(* Logix 5000 project; controller FV vendor 1 type 14 code 217 rev 31.11; software revision 31.00; part 42 of 63 *)
(* tags used below, declared in another part *)
   FV_B100 : INT[255];   // FV FLAGS
   FV_B100_0_1_OutputBit : BOOL;
   FV_N101 : INT[255];   // FV INT Fermentation control integer workspace
   FV_N110 : INT[255];   // FV DATA 0 CURRENT FV DATA
   FV_N12 : INT[255];   // SYS_PARMS System Parameter Fil e
   FV_SFile : INT[255];   // SLC Equivalent System File, So Original Code Can Remain
   FV_T102 : TIMER[20];
   FV_T4 : TIMER[10];
(* FV_Common, continued *)

ROUTINE FV_FV_ELAPSED_102   (* ladder *)
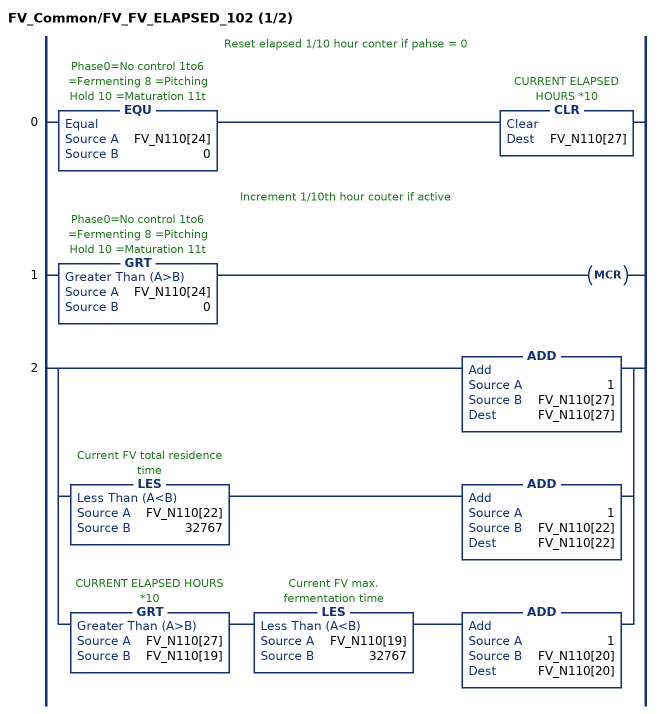
   // Reset elapsed 1/10 hour conter if pahse = 0
   0: EQU(FV_N110[24],0)CLR(FV_N110[27]);
   // Increment 1/10th hour couter if active
   1: GRT(FV_N110[24],0)MCR();
   2: [ADD(1,FV_N110[27],FV_N110[27]) ,LES(FV_N110[22],32767) ADD(1,FV_N110[22],FV_N110[22]) ,GRT(FV_N110[27],FV_N110[19]) LES(FV_N110[19],32767) ADD(1,FV_N110[20],FV_N110[20]) ];
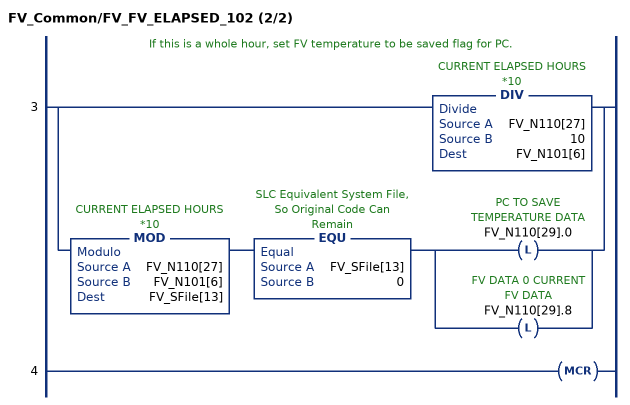
   // If this is a whole hour, set FV temperature to be saved flag for PC.
   3: [DIV(FV_N110[27],10,FV_N101[6]) ,MOD(FV_N110[27],FV_N101[6],FV_SFile[13]) EQU(FV_SFile[13],0) [OTL(FV_N110[29].0) ,OTL(FV_N110[29].8) ] ];
   4: MCR();
END_ROUTINE

ROUTINE FV_FV_MCP_100   (* ladder *)
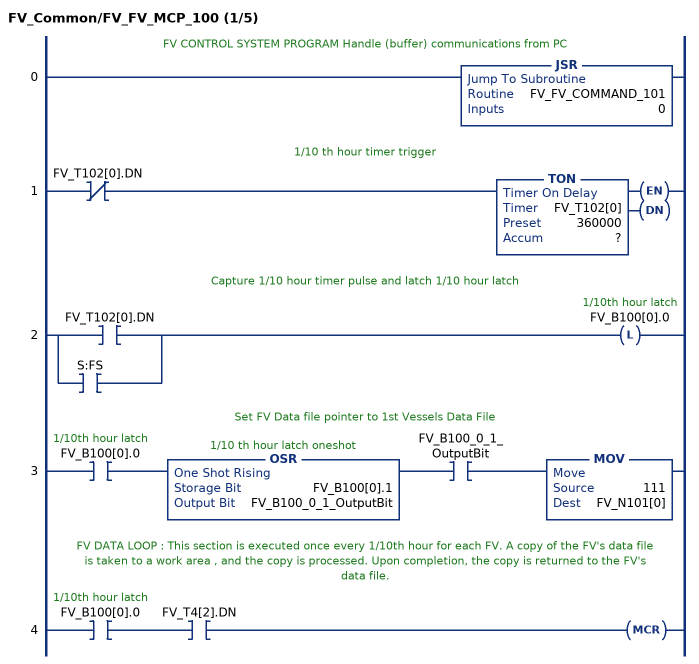
   // FV CONTROL SYSTEM PROGRAM Handle (buffer) communications from PC
   0: JSR(FV_FV_COMMAND_101,0);
   // 1/10 th hour timer trigger
   1: XIO(FV_T102[0].DN)TON(FV_T102[0],?,?);
   // Capture 1/10 hour timer pulse and latch 1/10 hour latch
   2: [XIC(FV_T102[0].DN) ,XIC(S:FS) ]OTL(FV_B100[0].0);
   // Set FV Data file pointer to 1st Vessels Data File
   3: XIC(FV_B100[0].0)OSR(FV_B100[0].1,FV_B100_0_1_OutputBit)XIC(FV_B100_0_1_OutputBit)MOV(111,FV_N101[0]);
   // FV DATA LOOP : This section is executed once every 1/10th hour for each FV. A copy of the FV's data file is taken to a work area , and the copy is processed. Upon completion, the copy is returned to the FV's data file.
   4: XIC(FV_B100[0].0)XIC(FV_T4[2].DN)MCR();
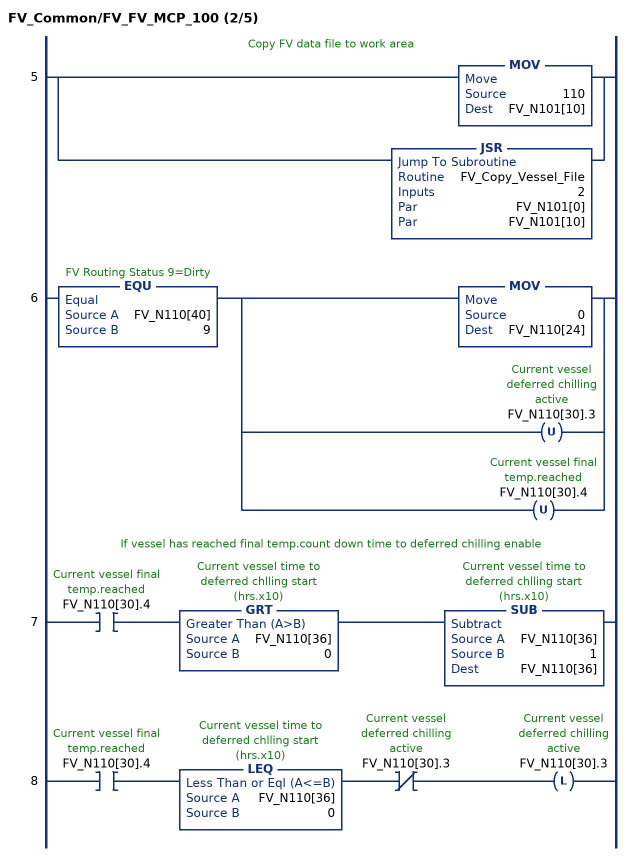
   // Copy FV data file to work area
   5: [MOV(110,FV_N101[10]) ,JSR(FV_Copy_Vessel_File,2,FV_N101[0],FV_N101[10]) ];
   6: EQU(FV_N110[40],9)[MOV(0,FV_N110[24]) ,OTU(FV_N110[30].3) ,OTU(FV_N110[30].4) ];
   // If vessel has reached final temp.count down time to deferred chilling enable
   7: XIC(FV_N110[30].4)GRT(FV_N110[36],0)SUB(FV_N110[36],1,FV_N110[36]);
   8: XIC(FV_N110[30].4)LEQ(FV_N110[36],0)XIO(FV_N110[30].3)OTL(FV_N110[30].3);
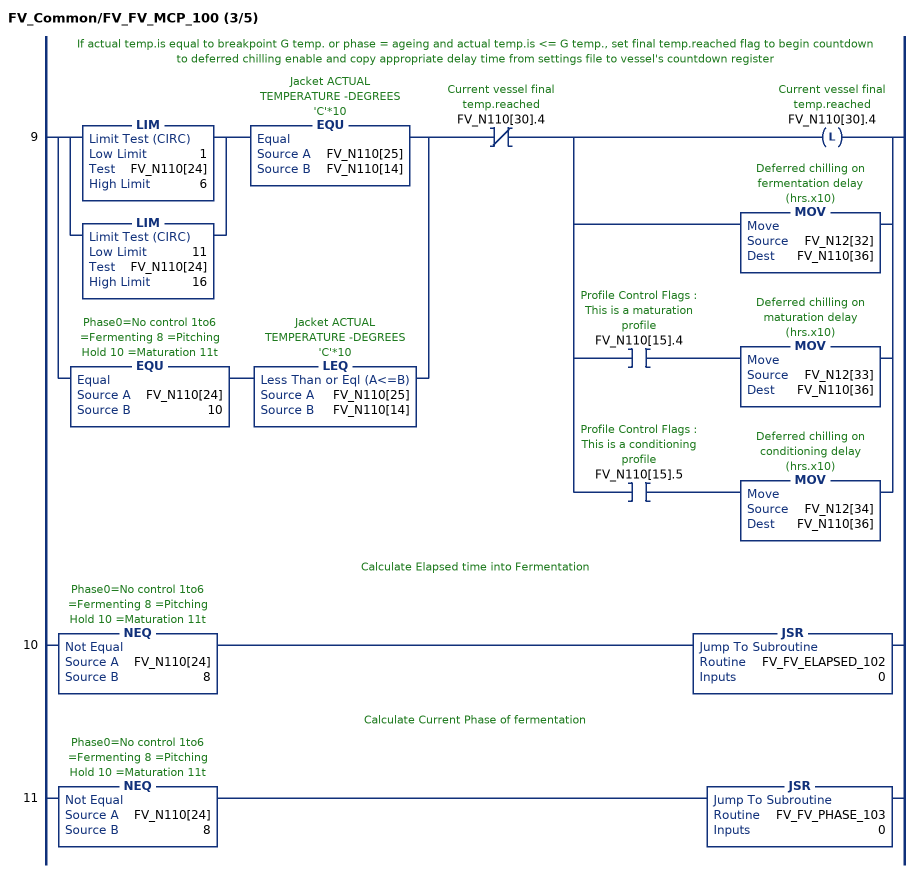
   // If actual temp.is equal to breakpoint G temp. or phase = ageing and actual temp.is <= G temp., set final temp.reached flag to begin countdown to deferred chilling enable and copy appropriate delay time from settings file to vessel's countdown register
   9: [[LIM(1,FV_N110[24],6) ,LIM(11,FV_N110[24],16) ] EQU(FV_N110[25],FV_N110[14]) ,EQU(FV_N110[24],10) LEQ(FV_N110[25],FV_N110[14]) ]XIO(FV_N110[30].4)[OTL(FV_N110[30].4) ,MOV(FV_N12[32],FV_N110[36]) ,XIC(FV_N110[15].4) MOV(FV_N12[33],FV_N110[36]) ,XIC(FV_N110[15].5) MOV(FV_N12[34],FV_N110[36]) ];
   // Calculate Elapsed time into Fermentation
   10: NEQ(FV_N110[24],8)JSR(FV_FV_ELAPSED_102,0);
   // Calculate Current Phase of fermentation
   11: NEQ(FV_N110[24],8)JSR(FV_FV_PHASE_103,0);
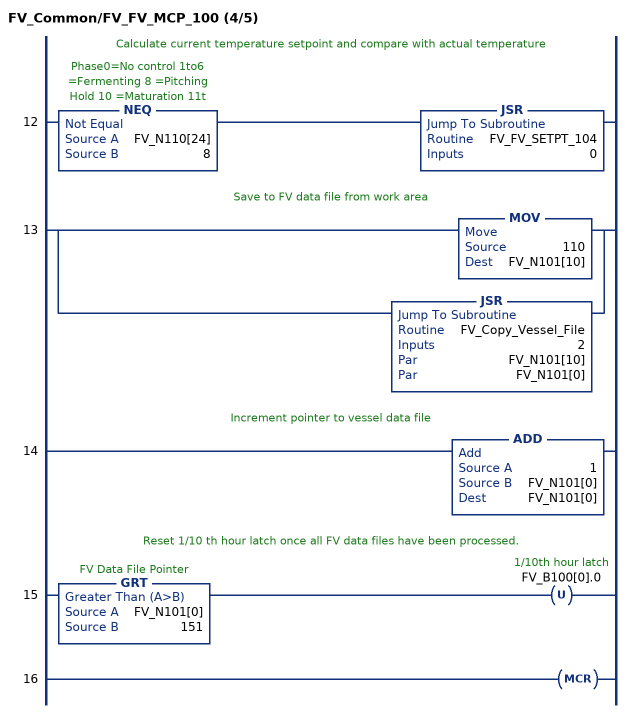
   // Calculate current temperature setpoint and compare with actual temperature
   12: NEQ(FV_N110[24],8)JSR(FV_FV_SETPT_104,0);
   // Save to FV data file from work area
   13: [MOV(110,FV_N101[10]) ,JSR(FV_Copy_Vessel_File,2,FV_N101[10],FV_N101[0]) ];
   // Increment pointer to vessel data file
   14: ADD(1,FV_N101[0],FV_N101[0]);
   // Reset 1/10 th hour latch once all FV data files have been processed.
   15: GRT(FV_N101[0],151)OTU(FV_B100[0].0);
   16: MCR();
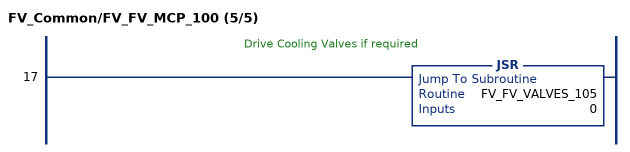
   // Drive Cooling Valves if required
   17: JSR(FV_FV_VALVES_105,0);
END_ROUTINE

ROUTINE FV_FV_PHASE_103   (* ladder *)
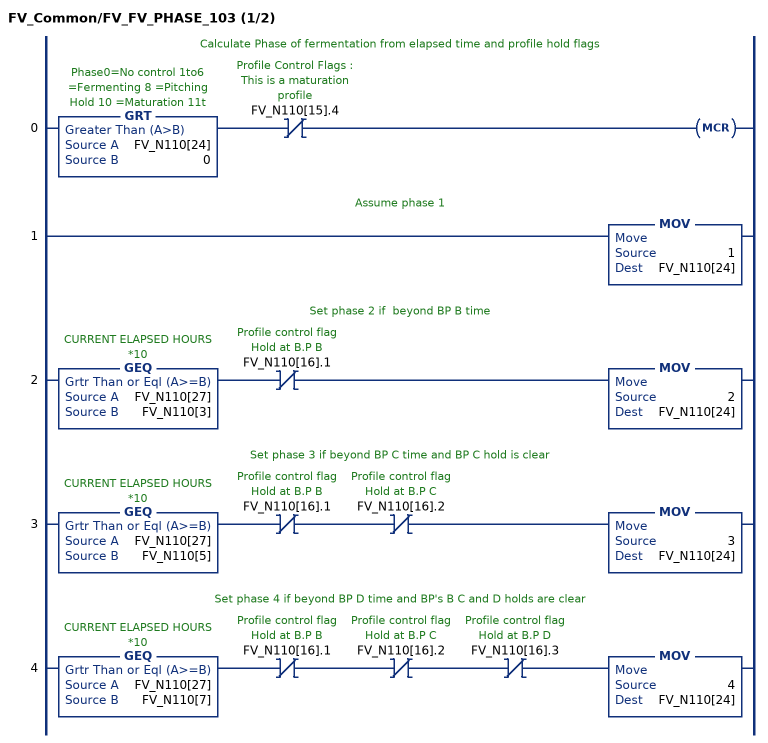
   // Calculate Phase of fermentation from elapsed time and profile hold flags
   0: GRT(FV_N110[24],0)XIO(FV_N110[15].4)MCR();
   // Assume phase 1
   1: MOV(1,FV_N110[24]);
   // Set phase 2 if  beyond BP B time
   2: GEQ(FV_N110[27],FV_N110[3])XIO(FV_N110[16].1)MOV(2,FV_N110[24]);
   // Set phase 3 if beyond BP C time and BP C hold is clear
   3: GEQ(FV_N110[27],FV_N110[5])XIO(FV_N110[16].1)XIO(FV_N110[16].2)MOV(3,FV_N110[24]);
   // Set phase 4 if beyond BP D time and BP's B C and D holds are clear
   4: GEQ(FV_N110[27],FV_N110[7])XIO(FV_N110[16].1)XIO(FV_N110[16].2)XIO(FV_N110[16].3)MOV(4,FV_N110[24]);
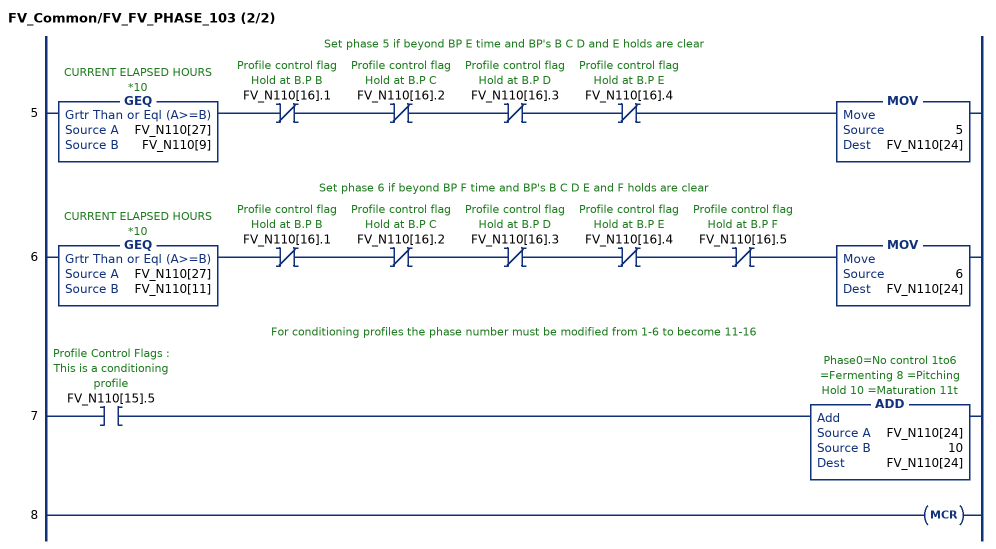
   // Set phase 5 if beyond BP E time and BP's B C D and E holds are clear
   5: GEQ(FV_N110[27],FV_N110[9])XIO(FV_N110[16].1)XIO(FV_N110[16].2)XIO(FV_N110[16].3)XIO(FV_N110[16].4)MOV(5,FV_N110[24]);
   // Set phase 6 if beyond BP F time and BP's B C D E and F holds are clear
   6: GEQ(FV_N110[27],FV_N110[11])XIO(FV_N110[16].1)XIO(FV_N110[16].2)XIO(FV_N110[16].3)XIO(FV_N110[16].4)XIO(FV_N110[16].5)MOV(6,FV_N110[24]);
   // For conditioning profiles the phase number must be modified from 1-6 to become 11-16
   7: XIC(FV_N110[15].5)ADD(FV_N110[24],10,FV_N110[24]);
   8: MCR();
END_ROUTINE

ROUTINE FV_FV_SETPT_104   (* ladder *)
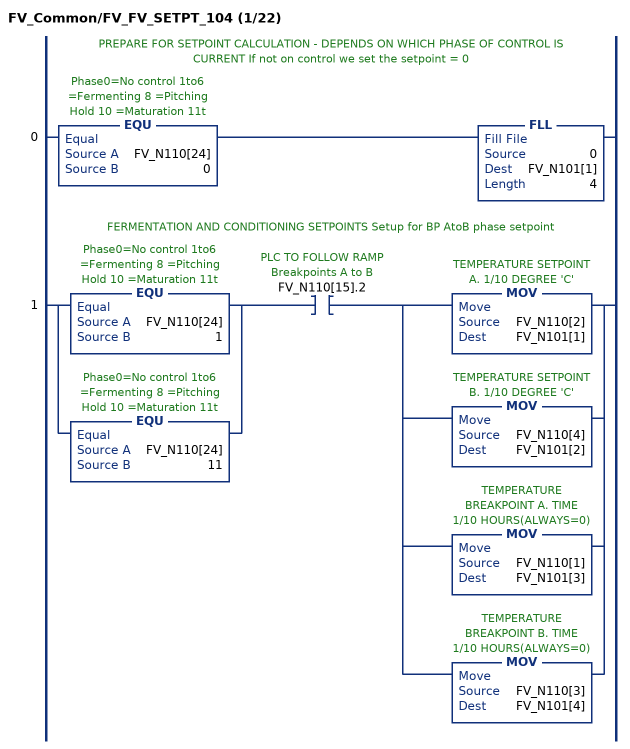
   // PREPARE FOR SETPOINT CALCULATION - DEPENDS ON WHICH PHASE OF CONTROL IS CURRENT If not on control we set the setpoint = 0
   0: EQU(FV_N110[24],0)FLL(0,FV_N101[1],4);
   // FERMENTATION AND CONDITIONING SETPOINTS Setup for BP AtoB phase setpoint
   1: [EQU(FV_N110[24],1) ,EQU(FV_N110[24],11) ]XIC(FV_N110[15].2)[MOV(FV_N110[2],FV_N101[1]) ,MOV(FV_N110[4],FV_N101[2]) ,MOV(FV_N110[1],FV_N101[3]) ,MOV(FV_N110[3],FV_N101[4]) ];
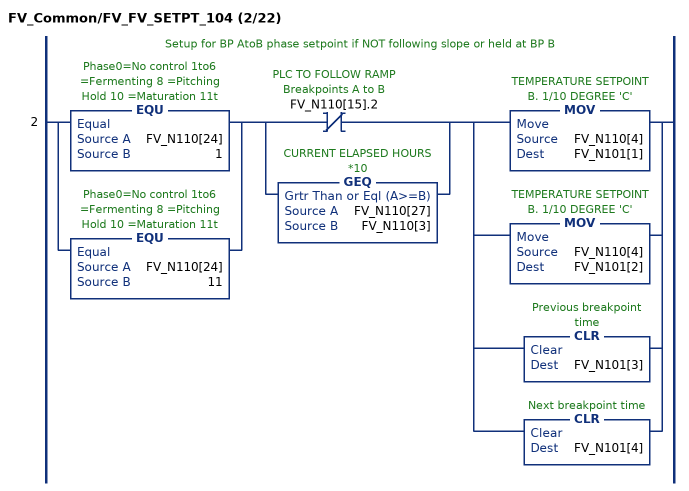
   // Setup for BP AtoB phase setpoint if NOT following slope or held at BP B
   2: [EQU(FV_N110[24],1) ,EQU(FV_N110[24],11) ][XIO(FV_N110[15].2) ,GEQ(FV_N110[27],FV_N110[3]) ][MOV(FV_N110[4],FV_N101[1]) ,MOV(FV_N110[4],FV_N101[2]) ,CLR(FV_N101[3]) ,CLR(FV_N101[4]) ];
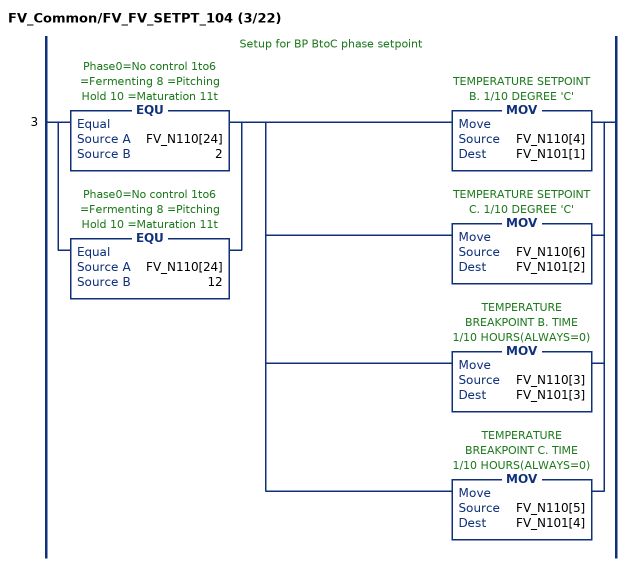
   // Setup for BP BtoC phase setpoint
   3: [EQU(FV_N110[24],2) ,EQU(FV_N110[24],12) ][MOV(FV_N110[4],FV_N101[1]) ,MOV(FV_N110[6],FV_N101[2]) ,MOV(FV_N110[3],FV_N101[3]) ,MOV(FV_N110[5],FV_N101[4]) ];
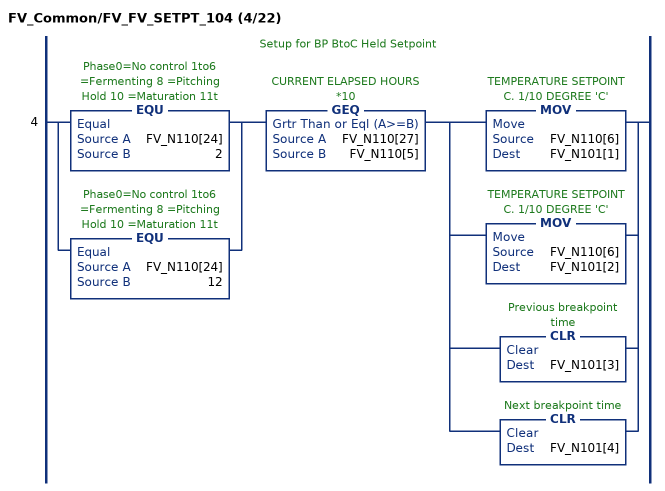
   // Setup for BP BtoC Held Setpoint
   4: [EQU(FV_N110[24],2) ,EQU(FV_N110[24],12) ]GEQ(FV_N110[27],FV_N110[5])[MOV(FV_N110[6],FV_N101[1]) ,MOV(FV_N110[6],FV_N101[2]) ,CLR(FV_N101[3]) ,CLR(FV_N101[4]) ];
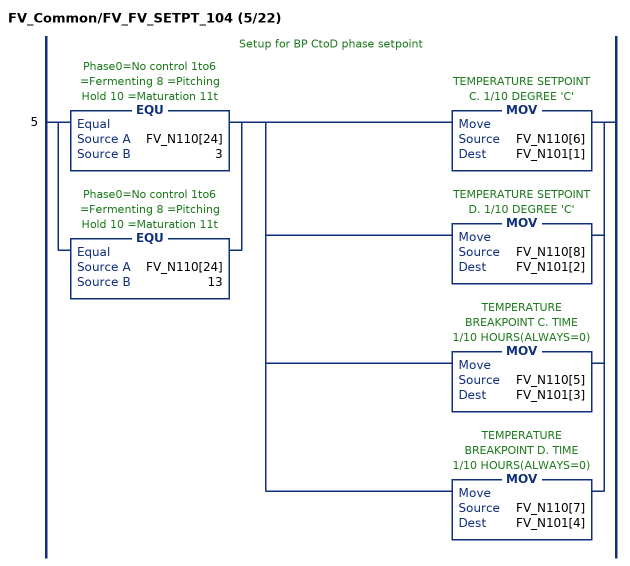
   // Setup for BP CtoD phase setpoint
   5: [EQU(FV_N110[24],3) ,EQU(FV_N110[24],13) ][MOV(FV_N110[6],FV_N101[1]) ,MOV(FV_N110[8],FV_N101[2]) ,MOV(FV_N110[5],FV_N101[3]) ,MOV(FV_N110[7],FV_N101[4]) ];
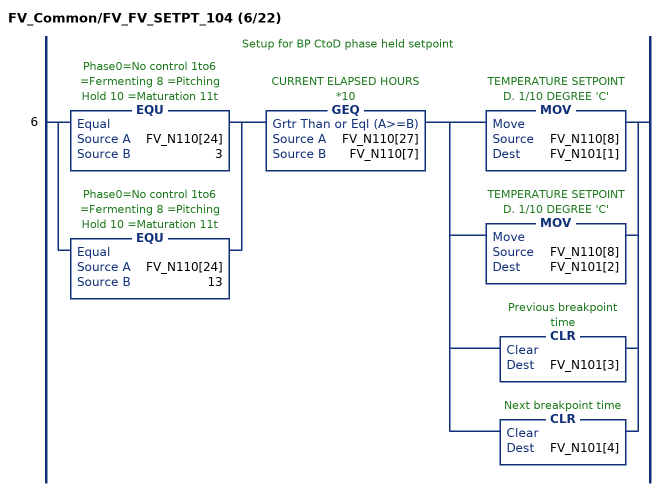
   // Setup for BP CtoD phase held setpoint
   6: [EQU(FV_N110[24],3) ,EQU(FV_N110[24],13) ]GEQ(FV_N110[27],FV_N110[7])[MOV(FV_N110[8],FV_N101[1]) ,MOV(FV_N110[8],FV_N101[2]) ,CLR(FV_N101[3]) ,CLR(FV_N101[4]) ];
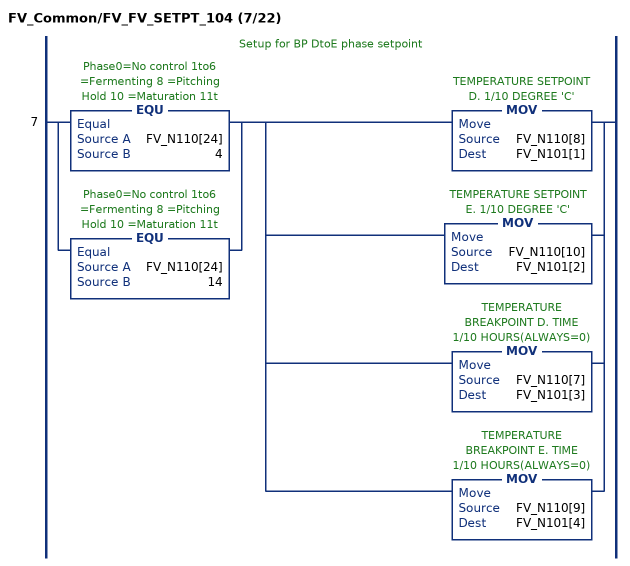
   // Setup for BP DtoE phase setpoint
   7: [EQU(FV_N110[24],4) ,EQU(FV_N110[24],14) ][MOV(FV_N110[8],FV_N101[1]) ,MOV(FV_N110[10],FV_N101[2]) ,MOV(FV_N110[7],FV_N101[3]) ,MOV(FV_N110[9],FV_N101[4]) ];
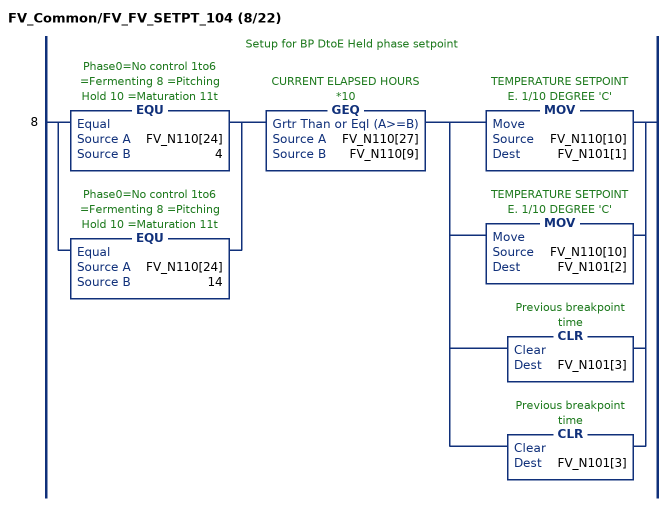
   // Setup for BP DtoE Held phase setpoint
   8: [EQU(FV_N110[24],4) ,EQU(FV_N110[24],14) ]GEQ(FV_N110[27],FV_N110[9])[MOV(FV_N110[10],FV_N101[1]) ,MOV(FV_N110[10],FV_N101[2]) ,CLR(FV_N101[3]) ,CLR(FV_N101[3]) ];
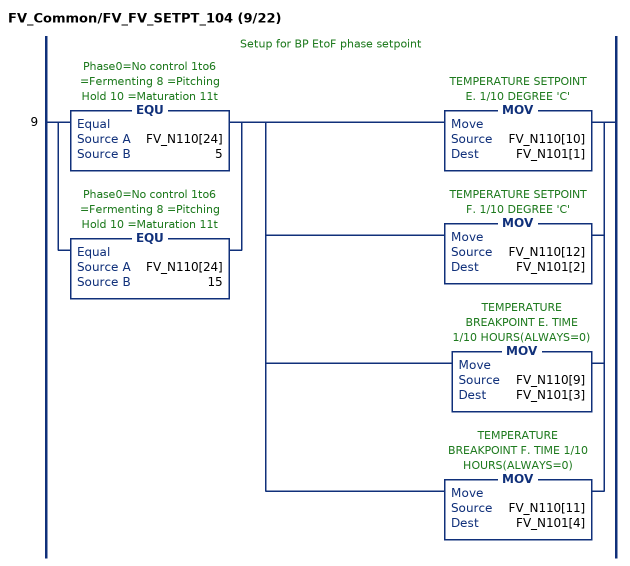
   // Setup for BP EtoF phase setpoint
   9: [EQU(FV_N110[24],5) ,EQU(FV_N110[24],15) ][MOV(FV_N110[10],FV_N101[1]) ,MOV(FV_N110[12],FV_N101[2]) ,MOV(FV_N110[9],FV_N101[3]) ,MOV(FV_N110[11],FV_N101[4]) ];
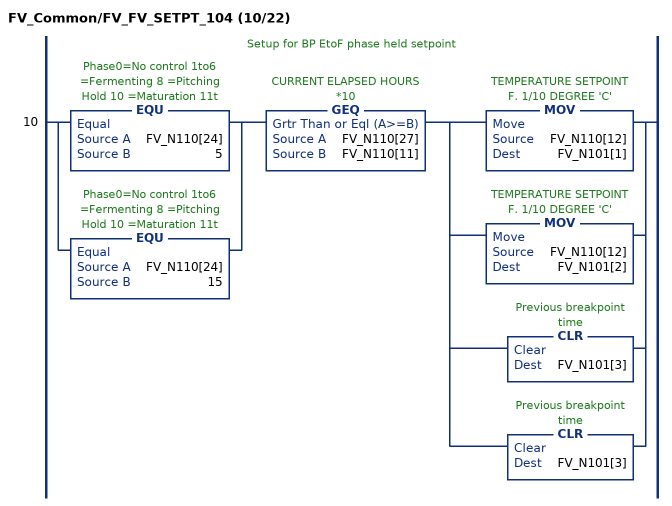
   // Setup for BP EtoF phase held setpoint
   10: [EQU(FV_N110[24],5) ,EQU(FV_N110[24],15) ]GEQ(FV_N110[27],FV_N110[11])[MOV(FV_N110[12],FV_N101[1]) ,MOV(FV_N110[12],FV_N101[2]) ,CLR(FV_N101[3]) ,CLR(FV_N101[3]) ];
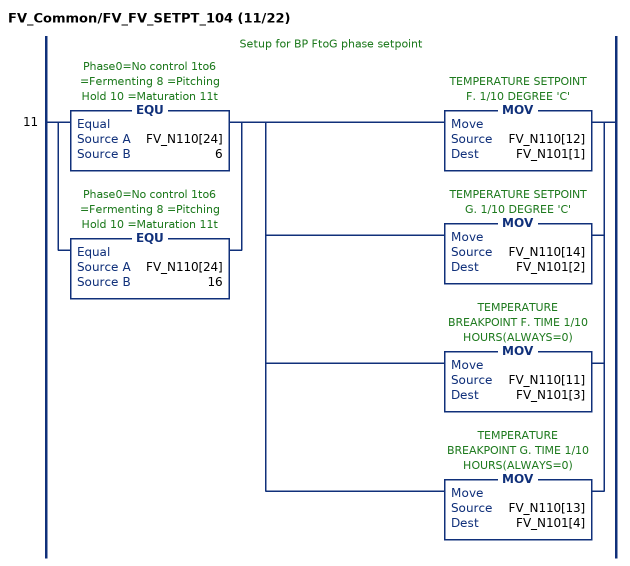
   // Setup for BP FtoG phase setpoint
   11: [EQU(FV_N110[24],6) ,EQU(FV_N110[24],16) ][MOV(FV_N110[12],FV_N101[1]) ,MOV(FV_N110[14],FV_N101[2]) ,MOV(FV_N110[11],FV_N101[3]) ,MOV(FV_N110[13],FV_N101[4]) ];
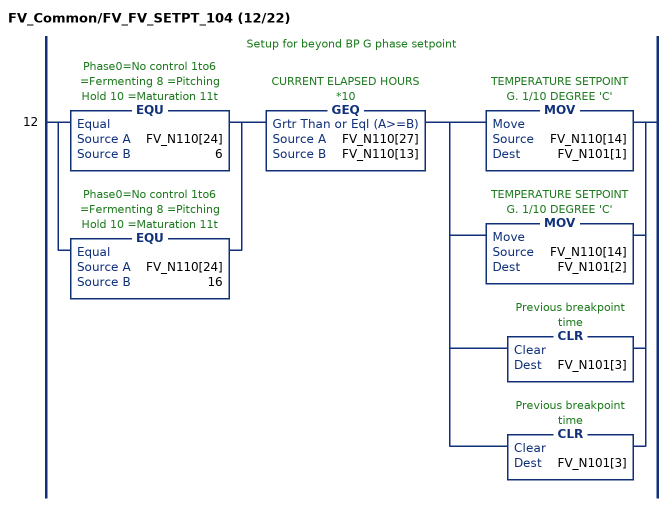
   // Setup for beyond BP G phase setpoint
   12: [EQU(FV_N110[24],6) ,EQU(FV_N110[24],16) ]GEQ(FV_N110[27],FV_N110[13])[MOV(FV_N110[14],FV_N101[1]) ,MOV(FV_N110[14],FV_N101[2]) ,CLR(FV_N101[3]) ,CLR(FV_N101[3]) ];
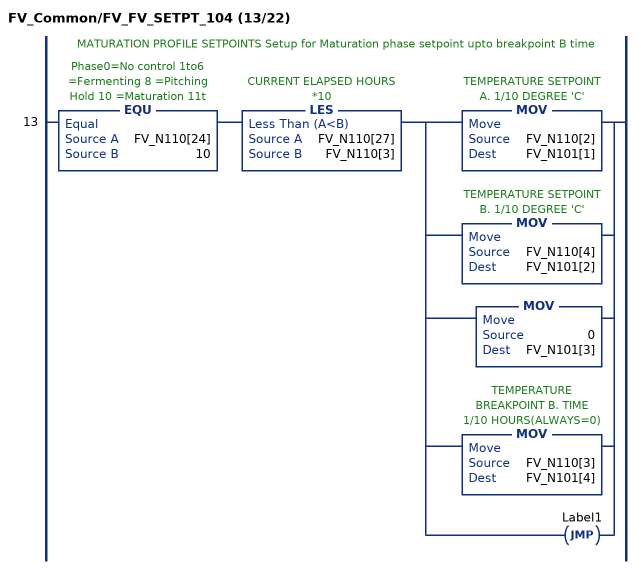
   // MATURATION PROFILE SETPOINTS Setup for Maturation phase setpoint upto breakpoint B time
   13: EQU(FV_N110[24],10)LES(FV_N110[27],FV_N110[3])[MOV(FV_N110[2],FV_N101[1]) ,MOV(FV_N110[4],FV_N101[2]) ,MOV(0,FV_N101[3]) ,MOV(FV_N110[3],FV_N101[4]) ,JMP(Label1) ];
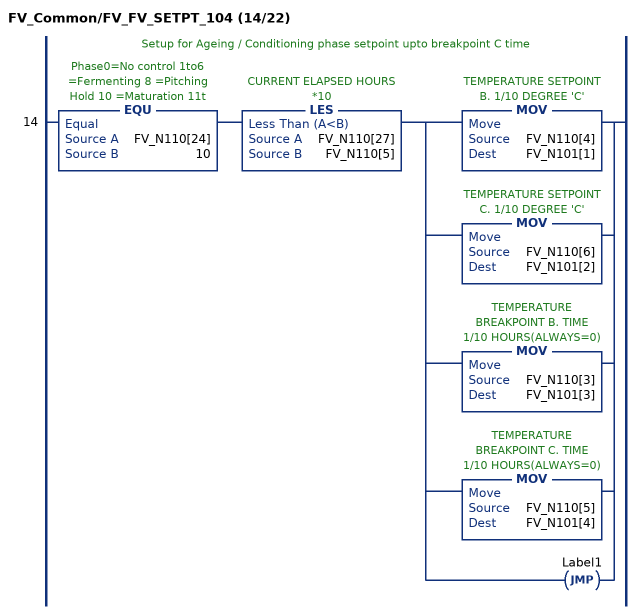
   // Setup for Ageing / Conditioning phase setpoint upto breakpoint C time
   14: EQU(FV_N110[24],10)LES(FV_N110[27],FV_N110[5])[MOV(FV_N110[4],FV_N101[1]) ,MOV(FV_N110[6],FV_N101[2]) ,MOV(FV_N110[3],FV_N101[3]) ,MOV(FV_N110[5],FV_N101[4]) ,JMP(Label1) ];
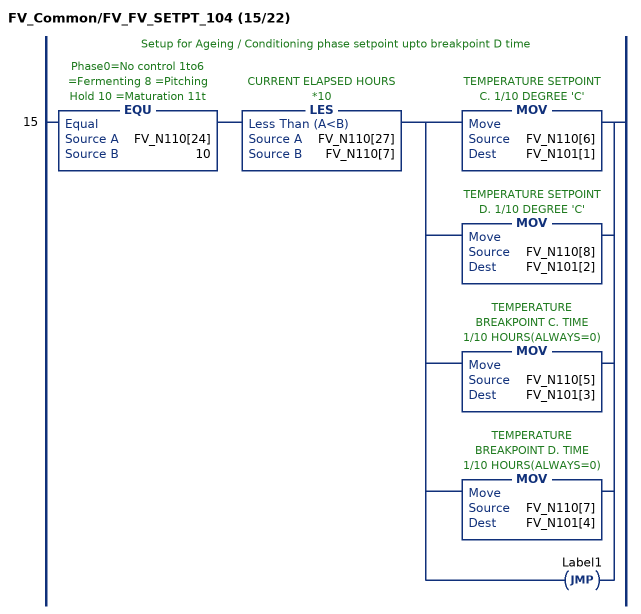
   // Setup for Ageing / Conditioning phase setpoint upto breakpoint D time
   15: EQU(FV_N110[24],10)LES(FV_N110[27],FV_N110[7])[MOV(FV_N110[6],FV_N101[1]) ,MOV(FV_N110[8],FV_N101[2]) ,MOV(FV_N110[5],FV_N101[3]) ,MOV(FV_N110[7],FV_N101[4]) ,JMP(Label1) ];
